REGION Network 157: Update the DAC for adjusting the VG2 voltage
   RUNG wire#powerrail
      { S7_Templates := "SrcType := Int" } LE_Contact(in1 := "STATO".stato_VOLTAGGIO_G2, in2 := 1150)
      { S7_Templates := "[SrcType := Int, DestType := Real]" } Convert(in := "STATO".stato_VOLTAGGIO_G2, out => "STATO_TMP".tmp_real_VG2)
      { S7_Templates := "SrcType := Real" } Mul(in1 := "STATO_TMP".tmp_real_VG2, in2 := 21.55, out => "STATO_TMP".tmp_real_VG2)
      { S7_Templates := "[SrcType := Real, DestType := DInt]" } Convert(in := "STATO_TMP".tmp_real_VG2, out => "STATO_TMP".tmp_adj_G2)
      { S7_Templates := "SrcType := DInt" } Mul(in1 := "STATO_TMP".tmp_adj_G2, in2 := "STATO".stato_adj_VG2, out => "STATO_TMP".tmp_adj_G2)
      { S7_Templates := "SrcType := DInt" } Div(in1 := "STATO_TMP".tmp_adj_G2, in2 := 1000, out => "dac_out_VG2")
   END_RUNG
   // the same network as SCL:
   IF "STATO".stato_VOLTAGGIO_G2 <= 1150 THEN
       "STATO_TMP".tmp_real_VG2 := INT_TO_REAL("STATO".stato_VOLTAGGIO_G2);
       "STATO_TMP".tmp_real_VG2 := "STATO_TMP".tmp_real_VG2 * 21.55;
       "STATO_TMP".tmp_adj_G2 := REAL_TO_DINT("STATO_TMP".tmp_real_VG2);
       "STATO_TMP".tmp_adj_G2 := "STATO_TMP".tmp_adj_G2 * "STATO".stato_adj_VG2;
       "dac_out_VG2" := "STATO_TMP".tmp_adj_G2 / 1000;
   END_IF;
END_REGION

REGION Network 158: Update the DAC for adjusting the VF voltage
   RUNG wire#powerrail
      { S7_Templates := "SrcType := Int" } LE_Contact(in1 := "STATO".stato_VOLTAGGIO_FILAMENTO, in2 := 8500)
      { S7_Templates := "[SrcType := Int, DestType := Real]" } Convert(in := "STATO".stato_VOLTAGGIO_FILAMENTO, out => "STATO_TMP".tmp_VFr)
      { S7_Templates := "SrcType := Real" } Div(in1 := "STATO_TMP".tmp_VFr, in2 := 1.0869, out => "STATO_TMP".tmp_VFr)
      { S7_Templates := "[SrcType := Real, DestType := Int]" } Convert(in := "STATO_TMP".tmp_VFr, out => "STATO_TMP".tmpVFi)
      { S7_Templates := "SrcType := DInt" } Mul(in1 := "STATO_TMP".tmpVFi, in2 := "STATO".stato_adj_VF, out => "STATO_TMP".tmp_adj_VF)
      { S7_Templates := "SrcType := DInt" } Div(in1 := "STATO_TMP".tmp_adj_VF, in2 := 1000, out => #dac_VF)
   END_RUNG
   // the same network as SCL:
   IF "STATO".stato_VOLTAGGIO_FILAMENTO <= 8500 THEN
       "STATO_TMP".tmp_VFr := INT_TO_REAL("STATO".stato_VOLTAGGIO_FILAMENTO);
       "STATO_TMP".tmp_VFr := "STATO_TMP".tmp_VFr / 1.0869;
       "STATO_TMP".tmpVFi := REAL_TO_INT("STATO_TMP".tmp_VFr);
       "STATO_TMP".tmp_adj_VF := "STATO_TMP".tmpVFi * "STATO".stato_adj_VF;
       #dac_VF := "STATO_TMP".tmp_adj_VF / 1000;
   END_IF;
END_REGION

REGION Network 159: Update the DAC for adjusting the VA voltage in CW
   // The voltage value must be below the threshold for CW mode.
   RUNG wire#powerrail
      Contact( "STATO".stato_MODO_CW )
      { S7_Templates := "SrcType := Int" } LE_Contact(in1 := "STATO".stato_ADJ_ANODICA_CW, in2 := "STATO".SOGLIA_VAcw)
      "REGOLA_ANODICA"(livello := "STATO".stato_ADJ_ANODICA_CW, uscita_dac => "dac_out_VA")
   END_RUNG
   // the same network as SCL:
   IF "STATO".stato_MODO_CW AND ("STATO".stato_ADJ_ANODICA_CW <= "STATO".SOGLIA_VAcw) THEN
       "REGOLA_ANODICA"(livello := "STATO".stato_ADJ_ANODICA_CW, uscita_dac => "dac_out_VA");
   END_IF;
END_REGION

REGION Network 160: Update the DAC for adjusting the VA voltage in Pulsed
   RUNG wire#powerrail
      Contact( "STATO".stato_MODO_PULSED )
      { S7_Templates := "SrcType := Int" } LE_Contact(in1 := "STATO".stato_ADJ_ANODICA_PULSED, in2 := 18000)
      "REGOLA_ANODICA"(livello := "STATO".stato_ADJ_ANODICA_PULSED, uscita_dac => "dac_out_VA")
   END_RUNG
   // the same network as SCL:
   IF "STATO".stato_MODO_PULSED AND ("STATO".stato_ADJ_ANODICA_PULSED <= 18000) THEN
       "REGOLA_ANODICA"(livello := "STATO".stato_ADJ_ANODICA_PULSED, uscita_dac => "dac_out_VA");
   END_IF;
END_REGION

REGION Network 161: Update the Reduced level
   RUNG wire#powerrail
      Contact( "STATO".controllo_setReduced )
      { S7_Templates := "SrcType := ???" } Mul(in1 := "STATO_TMP".tmp_Reduced, in2 := 10, out => "STATO".SogliaRidotta)
      Move(in := "STATO_TMP".tmp_Reduced, out1 => "STATO".stato_sogliaRIDOTTA)
      R_Coil( "STATO".controllo_setReduced )
   END_RUNG
   // the same network as SCL:
   IF "STATO".controllo_setReduced THEN
       "STATO".SogliaRidotta := "STATO_TMP".tmp_Reduced * 10;
       "STATO".stato_sogliaRIDOTTA := "STATO_TMP".tmp_Reduced;
       "STATO".controllo_setReduced := FALSE;
   END_IF;
END_REGION

REGION Network 162: Update the power levels for display panel
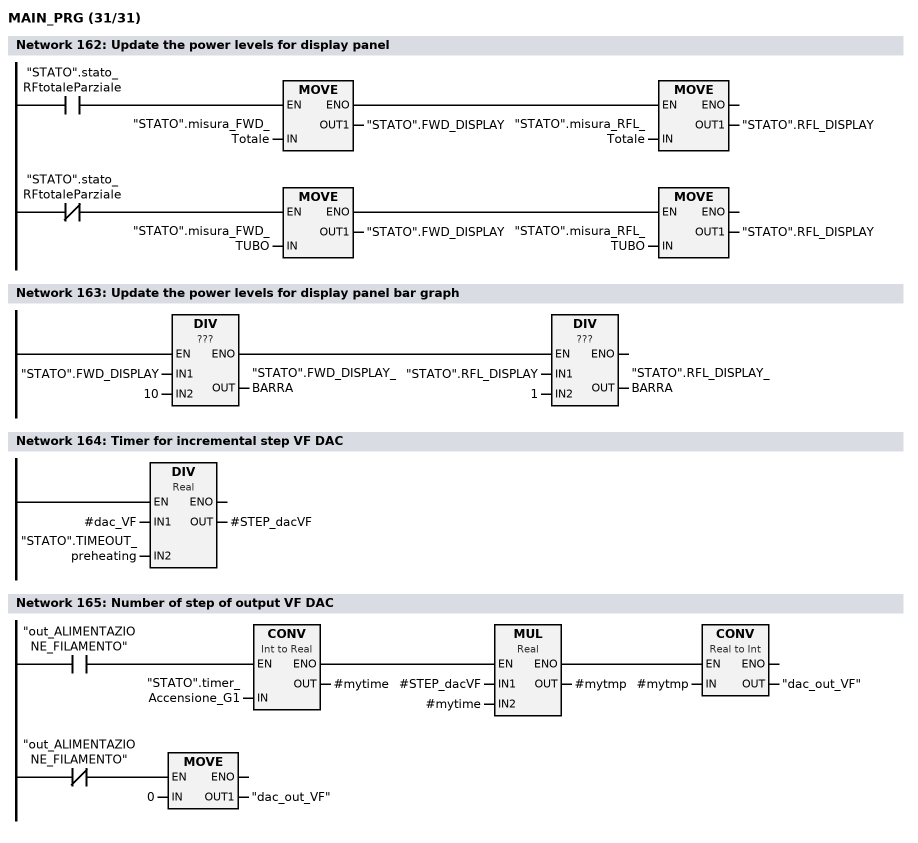
   RUNG wire#powerrail
      Contact( "STATO".stato_RFtotaleParziale )
      Move(in := "STATO".misura_FWD_Totale, out1 => "STATO".FWD_DISPLAY)
      Move(in := "STATO".misura_RFL_Totale, out1 => "STATO".RFL_DISPLAY)
   END_RUNG
   RUNG wire#powerrail
      I_Contact( "STATO".stato_RFtotaleParziale )
      Move(in := "STATO".misura_FWD_TUBO, out1 => "STATO".FWD_DISPLAY)
      Move(in := "STATO".misura_RFL_TUBO, out1 => "STATO".RFL_DISPLAY)
   END_RUNG
   // the same network as SCL:
   IF "STATO".stato_RFtotaleParziale THEN
       "STATO".FWD_DISPLAY := "STATO".misura_FWD_Totale;
       "STATO".RFL_DISPLAY := "STATO".misura_RFL_Totale;
   END_IF;
   IF NOT "STATO".stato_RFtotaleParziale THEN
       "STATO".FWD_DISPLAY := "STATO".misura_FWD_TUBO;
       "STATO".RFL_DISPLAY := "STATO".misura_RFL_TUBO;
   END_IF;
END_REGION

REGION Network 163: Update the power levels for display panel bar graph
   RUNG wire#powerrail
      { S7_Templates := "SrcType := ???" } Div(in1 := "STATO".FWD_DISPLAY, in2 := 10, out => "STATO".FWD_DISPLAY_BARRA)
      { S7_Templates := "SrcType := ???" } Div(in1 := "STATO".RFL_DISPLAY, in2 := 1, out => "STATO".RFL_DISPLAY_BARRA)
   END_RUNG
   // the same network as SCL:
   "STATO".FWD_DISPLAY_BARRA := "STATO".FWD_DISPLAY / 10;
   "STATO".RFL_DISPLAY_BARRA := "STATO".RFL_DISPLAY / 1;
END_REGION

REGION Network 164: Timer for incremental step VF DAC
   RUNG wire#powerrail
      { S7_Templates := "SrcType := Real" } Div(in1 := #dac_VF, in2 := "STATO".TIMEOUT_preheating, out => #STEP_dacVF)
   END_RUNG
   // the same network as SCL:
   #STEP_dacVF := #dac_VF / "STATO".TIMEOUT_preheating;
END_REGION

REGION Network 165: Number of step of output VF DAC
   RUNG wire#powerrail
      Contact( "out_ALIMENTAZIONE_FILAMENTO" )
      { S7_Templates := "[SrcType := Int, DestType := Real]" } Convert(in := "STATO".timer_Accensione_G1, out => #mytime)
      { S7_Templates := "SrcType := Real" } Mul(in1 := #STEP_dacVF, in2 := #mytime, out => #mytmp)
      { S7_Templates := "[SrcType := Real, DestType := Int]" } Convert(in := #mytmp, out => "dac_out_VF")
   END_RUNG
   RUNG wire#powerrail
      I_Contact( "out_ALIMENTAZIONE_FILAMENTO" )
      Move(in := 0, out1 => "dac_out_VF")
   END_RUNG
   // the same network as SCL:
   IF "out_ALIMENTAZIONE_FILAMENTO" THEN
       #mytime := INT_TO_REAL("STATO".timer_Accensione_G1);
       #mytmp := #STEP_dacVF * #mytime;
       "dac_out_VF" := REAL_TO_INT(#mytmp);
   END_IF;
   IF NOT "out_ALIMENTAZIONE_FILAMENTO" THEN "dac_out_VF" := 0; END_IF;
END_REGION
END_FUNCTION_BLOCK

FUNCTION "MISURE_ANALOGICHE" : Void   // FC1, LAD
TITLE = LETTURE ANALOGICHE DALL'ADC E DAL FLUSSOMETRO
{ S7_Optimized_Access := 'FALSE' }
VERSION : 0.1
   VAR_TEMP   // added for the SCL form of the ladder/FBD networks
      _w1 : Bool;
      _w2 : Bool;
      _w3 : Bool;
   END_VAR
BEGIN

REGION Network 1: MISURA TEMPERATURA LQD IN SS (1) bloccato
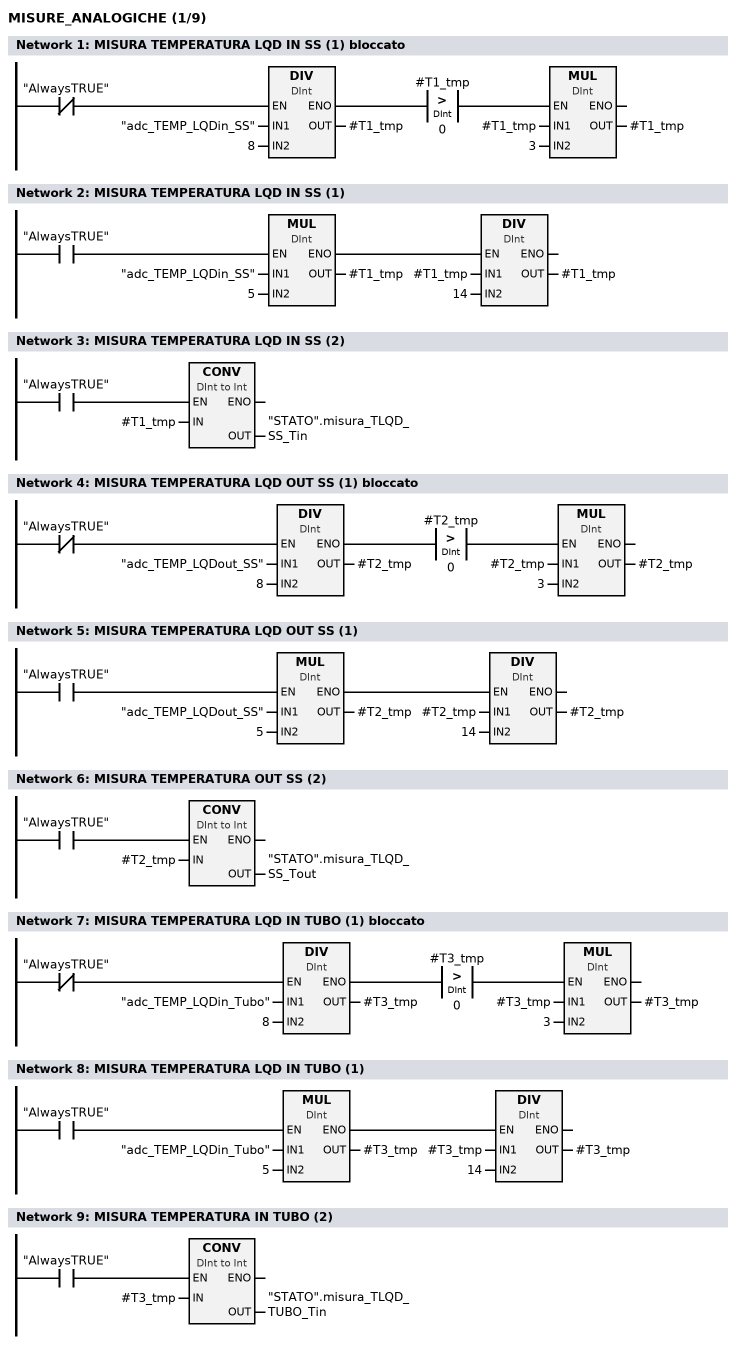
   RUNG wire#powerrail
      I_Contact( "AlwaysTRUE" )
      { S7_Templates := "SrcType := DInt" } Div(in1 := "adc_TEMP_LQDin_SS", in2 := 8, out => #T1_tmp)
      { S7_Templates := "SrcType := DInt" } GT_Contact(in1 := #T1_tmp, in2 := 0)
      { S7_Templates := "SrcType := DInt" } Mul(in1 := #T1_tmp, in2 := 3, out => #T1_tmp)
   END_RUNG
   // the same network as SCL:
   IF NOT "AlwaysTRUE" THEN #T1_tmp := "adc_TEMP_LQDin_SS" / 8; END_IF;
   IF NOT "AlwaysTRUE" AND (#T1_tmp > 0) THEN #T1_tmp := #T1_tmp * 3; END_IF;
END_REGION

REGION Network 2: MISURA TEMPERATURA LQD IN SS (1)
   RUNG wire#powerrail
      Contact( "AlwaysTRUE" )
      { S7_Templates := "SrcType := DInt" } Mul(in1 := "adc_TEMP_LQDin_SS", in2 := 5, out => #T1_tmp)
      { S7_Templates := "SrcType := DInt" } Div(in1 := #T1_tmp, in2 := 14, out => #T1_tmp)
   END_RUNG
   // the same network as SCL:
   IF "AlwaysTRUE" THEN
       #T1_tmp := "adc_TEMP_LQDin_SS" * 5;
       #T1_tmp := #T1_tmp / 14;
   END_IF;
END_REGION

REGION Network 3: MISURA TEMPERATURA LQD IN SS (2)
   RUNG wire#powerrail
      Contact( "AlwaysTRUE" )
      { S7_Templates := "[SrcType := DInt, DestType := Int]" } Convert(in := #T1_tmp, out => "STATO".misura_TLQD_SS_Tin)
   END_RUNG
   // the same network as SCL:
   IF "AlwaysTRUE" THEN "STATO".misura_TLQD_SS_Tin := DINT_TO_INT(#T1_tmp); END_IF;
END_REGION

REGION Network 4: MISURA TEMPERATURA LQD OUT SS (1) bloccato
   RUNG wire#powerrail
      I_Contact( "AlwaysTRUE" )
      { S7_Templates := "SrcType := DInt" } Div(in1 := "adc_TEMP_LQDout_SS", in2 := 8, out => #T2_tmp)
      { S7_Templates := "SrcType := DInt" } GT_Contact(in1 := #T2_tmp, in2 := 0)
      { S7_Templates := "SrcType := DInt" } Mul(in1 := #T2_tmp, in2 := 3, out => #T2_tmp)
   END_RUNG
   // the same network as SCL:
   IF NOT "AlwaysTRUE" THEN #T2_tmp := "adc_TEMP_LQDout_SS" / 8; END_IF;
   IF NOT "AlwaysTRUE" AND (#T2_tmp > 0) THEN #T2_tmp := #T2_tmp * 3; END_IF;
END_REGION

REGION Network 5: MISURA TEMPERATURA LQD OUT SS (1)
   RUNG wire#powerrail
      Contact( "AlwaysTRUE" )
      { S7_Templates := "SrcType := DInt" } Mul(in1 := "adc_TEMP_LQDout_SS", in2 := 5, out => #T2_tmp)
      { S7_Templates := "SrcType := DInt" } Div(in1 := #T2_tmp, in2 := 14, out => #T2_tmp)
   END_RUNG
   // the same network as SCL:
   IF "AlwaysTRUE" THEN
       #T2_tmp := "adc_TEMP_LQDout_SS" * 5;
       #T2_tmp := #T2_tmp / 14;
   END_IF;
END_REGION

REGION Network 6: MISURA TEMPERATURA OUT SS (2)
   RUNG wire#powerrail
      Contact( "AlwaysTRUE" )
      { S7_Templates := "[SrcType := DInt, DestType := Int]" } Convert(in := #T2_tmp, out => "STATO".misura_TLQD_SS_Tout)
   END_RUNG
   // the same network as SCL:
   IF "AlwaysTRUE" THEN "STATO".misura_TLQD_SS_Tout := DINT_TO_INT(#T2_tmp); END_IF;
END_REGION

REGION Network 7: MISURA TEMPERATURA LQD IN TUBO (1) bloccato
   RUNG wire#powerrail
      I_Contact( "AlwaysTRUE" )
      { S7_Templates := "SrcType := DInt" } Div(in1 := "adc_TEMP_LQDin_Tubo", in2 := 8, out => #T3_tmp)
      { S7_Templates := "SrcType := DInt" } GT_Contact(in1 := #T3_tmp, in2 := 0)
      { S7_Templates := "SrcType := DInt" } Mul(in1 := #T3_tmp, in2 := 3, out => #T3_tmp)
   END_RUNG
   // the same network as SCL:
   IF NOT "AlwaysTRUE" THEN #T3_tmp := "adc_TEMP_LQDin_Tubo" / 8; END_IF;
   IF NOT "AlwaysTRUE" AND (#T3_tmp > 0) THEN #T3_tmp := #T3_tmp * 3; END_IF;
END_REGION

REGION Network 8: MISURA TEMPERATURA LQD IN TUBO (1)
   RUNG wire#powerrail
      Contact( "AlwaysTRUE" )
      { S7_Templates := "SrcType := DInt" } Mul(in1 := "adc_TEMP_LQDin_Tubo", in2 := 5, out => #T3_tmp)
      { S7_Templates := "SrcType := DInt" } Div(in1 := #T3_tmp, in2 := 14, out => #T3_tmp)
   END_RUNG
   // the same network as SCL:
   IF "AlwaysTRUE" THEN
       #T3_tmp := "adc_TEMP_LQDin_Tubo" * 5;
       #T3_tmp := #T3_tmp / 14;
   END_IF;
END_REGION

REGION Network 9: MISURA TEMPERATURA IN TUBO (2)
   RUNG wire#powerrail
      Contact( "AlwaysTRUE" )
      { S7_Templates := "[SrcType := DInt, DestType := Int]" } Convert(in := #T3_tmp, out => "STATO".misura_TLQD_TUBO_Tin)
   END_RUNG
   // the same network as SCL:
   IF "AlwaysTRUE" THEN "STATO".misura_TLQD_TUBO_Tin := DINT_TO_INT(#T3_tmp); END_IF;
END_REGION

REGION Network 10: MISURA TEMPERATURA LQD OUT TUBO (1) bloccato
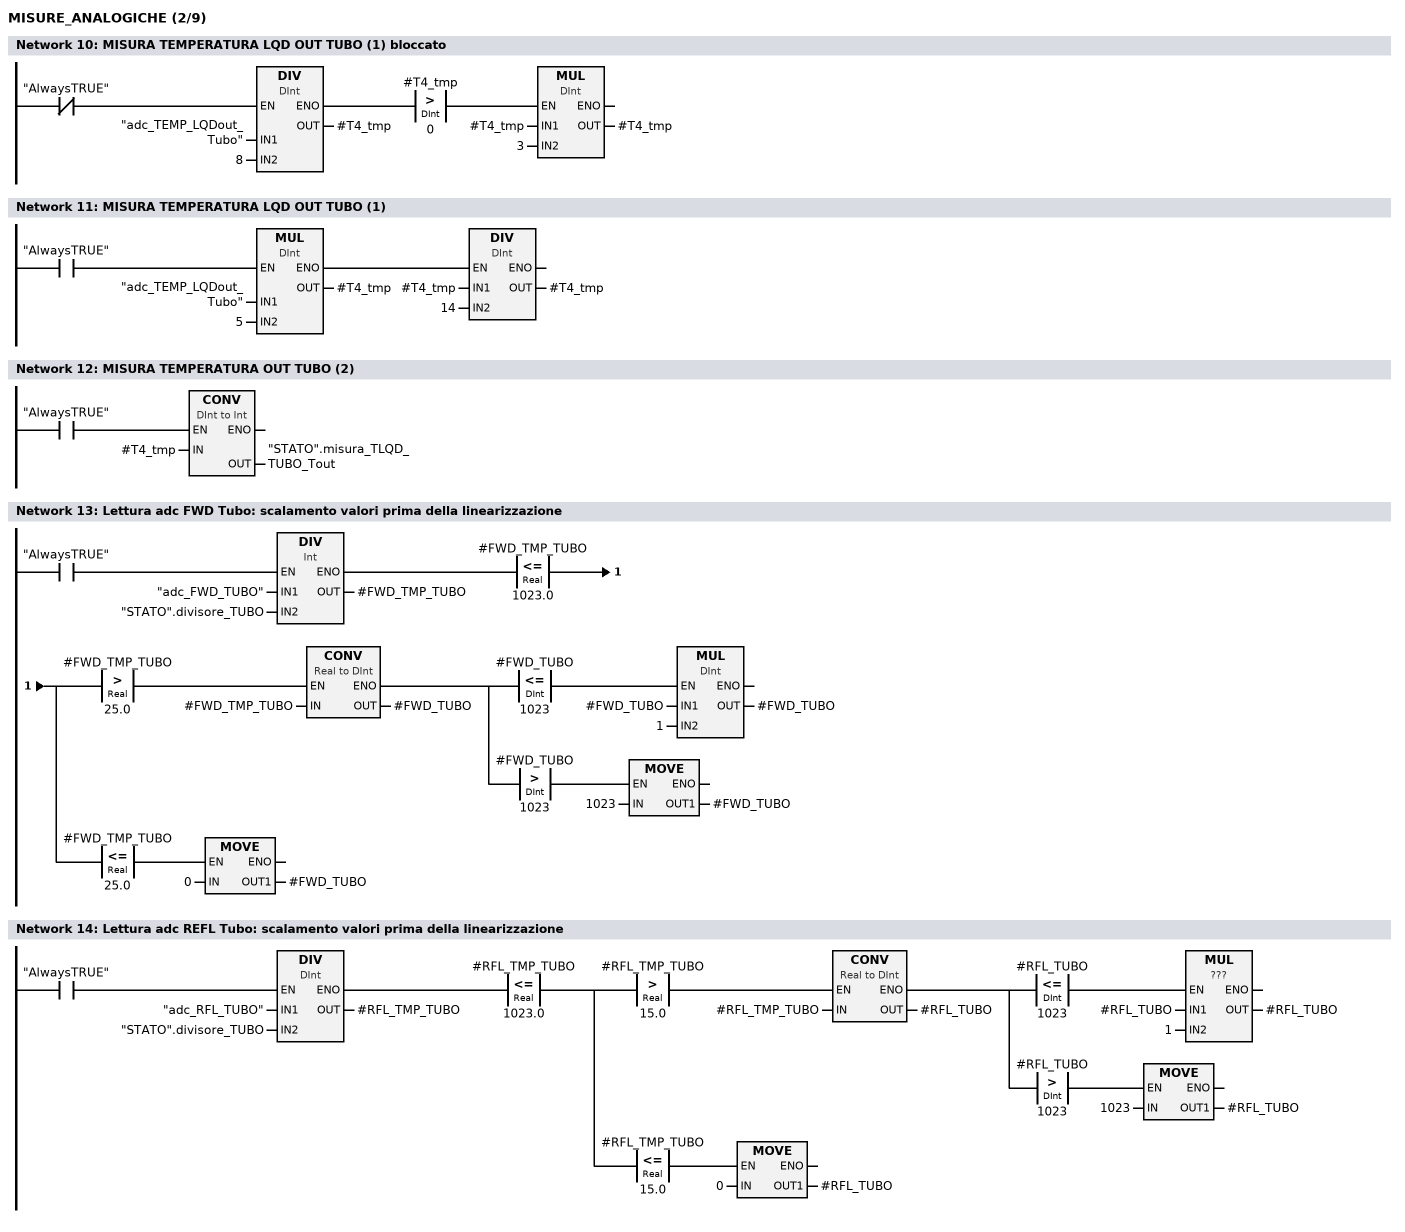
   RUNG wire#powerrail
      I_Contact( "AlwaysTRUE" )
      { S7_Templates := "SrcType := DInt" } Div(in1 := "adc_TEMP_LQDout_Tubo", in2 := 8, out => #T4_tmp)
      { S7_Templates := "SrcType := DInt" } GT_Contact(in1 := #T4_tmp, in2 := 0)
      { S7_Templates := "SrcType := DInt" } Mul(in1 := #T4_tmp, in2 := 3, out => #T4_tmp)
   END_RUNG
   // the same network as SCL:
   IF NOT "AlwaysTRUE" THEN #T4_tmp := "adc_TEMP_LQDout_Tubo" / 8; END_IF;
   IF NOT "AlwaysTRUE" AND (#T4_tmp > 0) THEN #T4_tmp := #T4_tmp * 3; END_IF;
END_REGION

REGION Network 11: MISURA TEMPERATURA LQD OUT TUBO (1)
   RUNG wire#powerrail
      Contact( "AlwaysTRUE" )
      { S7_Templates := "SrcType := DInt" } Mul(in1 := "adc_TEMP_LQDout_Tubo", in2 := 5, out => #T4_tmp)
      { S7_Templates := "SrcType := DInt" } Div(in1 := #T4_tmp, in2 := 14, out => #T4_tmp)
   END_RUNG
   // the same network as SCL:
   IF "AlwaysTRUE" THEN
       #T4_tmp := "adc_TEMP_LQDout_Tubo" * 5;
       #T4_tmp := #T4_tmp / 14;
   END_IF;
END_REGION

REGION Network 12: MISURA TEMPERATURA OUT TUBO (2)
   RUNG wire#powerrail
      Contact( "AlwaysTRUE" )
      { S7_Templates := "[SrcType := DInt, DestType := Int]" } Convert(in := #T4_tmp, out => "STATO".misura_TLQD_TUBO_Tout)
   END_RUNG
   // the same network as SCL:
   IF "AlwaysTRUE" THEN "STATO".misura_TLQD_TUBO_Tout := DINT_TO_INT(#T4_tmp); END_IF;
END_REGION

REGION Network 13: Lettura adc FWD Tubo: scalamento valori prima della linearizzazione
   RUNG wire#powerrail
      Contact( "AlwaysTRUE" )
      { S7_Templates := "SrcType := Int" } Div(in1 := "adc_FWD_TUBO", in2 := "STATO".divisore_TUBO, out => #FWD_TMP_TUBO)
      { S7_Templates := "SrcType := Real" } LE_Contact(in1 := #FWD_TMP_TUBO, in2 := 1023.0)
      wire#w1
      { S7_Templates := "SrcType := Real" } GT_Contact(in1 := #FWD_TMP_TUBO, in2 := 25.0)
      { S7_Templates := "[SrcType := Real, DestType := DInt]" } Convert(in := #FWD_TMP_TUBO, out => #FWD_TUBO)
      wire#w2
      { S7_Templates := "SrcType := DInt" } LE_Contact(in1 := #FWD_TUBO, in2 := 1023)
      { S7_Templates := "SrcType := DInt" } Mul(in1 := #FWD_TUBO, in2 := 1, out => #FWD_TUBO)
   END_RUNG
   RUNG wire#w2
      { S7_Templates := "SrcType := DInt" } GT_Contact(in1 := #FWD_TUBO, in2 := 1023)
      Move(in := 1023, out1 => #FWD_TUBO)
   END_RUNG
   RUNG wire#w1
      { S7_Templates := "SrcType := Real" } LE_Contact(in1 := #FWD_TMP_TUBO, in2 := 25.0)
      Move(in := 0, out1 => #FWD_TUBO)
   END_RUNG
   // the same network as SCL:
   IF "AlwaysTRUE" THEN #FWD_TMP_TUBO := "adc_FWD_TUBO" / "STATO".divisore_TUBO; END_IF;
   #_w1 := "AlwaysTRUE" AND (#FWD_TMP_TUBO <= 1023.0);
   #_w2 := #_w1 AND (#FWD_TMP_TUBO > 25.0);
   IF #_w2 THEN #FWD_TUBO := REAL_TO_DINT(#FWD_TMP_TUBO); END_IF;
   IF #_w2 AND (#FWD_TUBO <= 1023) THEN #FWD_TUBO := #FWD_TUBO * 1; END_IF;
   IF #_w2 AND (#FWD_TUBO > 1023) THEN #FWD_TUBO := 1023; END_IF;
   IF #_w1 AND (#FWD_TMP_TUBO <= 25.0) THEN #FWD_TUBO := 0; END_IF;
END_REGION

REGION Network 14: Lettura adc REFL Tubo: scalamento valori prima della linearizzazione
   RUNG wire#powerrail
      Contact( "AlwaysTRUE" )
      { S7_Templates := "SrcType := DInt" } Div(in1 := "adc_RFL_TUBO", in2 := "STATO".divisore_TUBO, out => #RFL_TMP_TUBO)
      { S7_Templates := "SrcType := Real" } LE_Contact(in1 := #RFL_TMP_TUBO, in2 := 1023.0)
      wire#w1
      { S7_Templates := "SrcType := Real" } GT_Contact(in1 := #RFL_TMP_TUBO, in2 := 15.0)
      { S7_Templates := "[SrcType := Real, DestType := DInt]" } Convert(in := #RFL_TMP_TUBO, out => #RFL_TUBO)
      wire#w2
      { S7_Templates := "SrcType := DInt" } LE_Contact(in1 := #RFL_TUBO, in2 := 1023)
      { S7_Templates := "SrcType := ???" } Mul(in1 := #RFL_TUBO, in2 := 1, out => #RFL_TUBO)
   END_RUNG
   RUNG wire#w2
      { S7_Templates := "SrcType := DInt" } GT_Contact(in1 := #RFL_TUBO, in2 := 1023)
      Move(in := 1023, out1 => #RFL_TUBO)
   END_RUNG
   RUNG wire#w1
      { S7_Templates := "SrcType := Real" } LE_Contact(in1 := #RFL_TMP_TUBO, in2 := 15.0)
      Move(in := 0, out1 => #RFL_TUBO)
   END_RUNG
   // the same network as SCL:
   IF "AlwaysTRUE" THEN #RFL_TMP_TUBO := "adc_RFL_TUBO" / "STATO".divisore_TUBO; END_IF;
   #_w1 := "AlwaysTRUE" AND (#RFL_TMP_TUBO <= 1023.0);
   #_w2 := #_w1 AND (#RFL_TMP_TUBO > 15.0);
   IF #_w2 THEN #RFL_TUBO := REAL_TO_DINT(#RFL_TMP_TUBO); END_IF;
   IF #_w2 AND (#RFL_TUBO <= 1023) THEN #RFL_TUBO := #RFL_TUBO * 1; END_IF;
   IF #_w2 AND (#RFL_TUBO > 1023) THEN #RFL_TUBO := 1023; END_IF;
   IF #_w1 AND (#RFL_TMP_TUBO <= 15.0) THEN #RFL_TUBO := 0; END_IF;
END_REGION

REGION Network 15: Lettura adc FWD Stato Solido: scalamento valori prima della linearizzazione
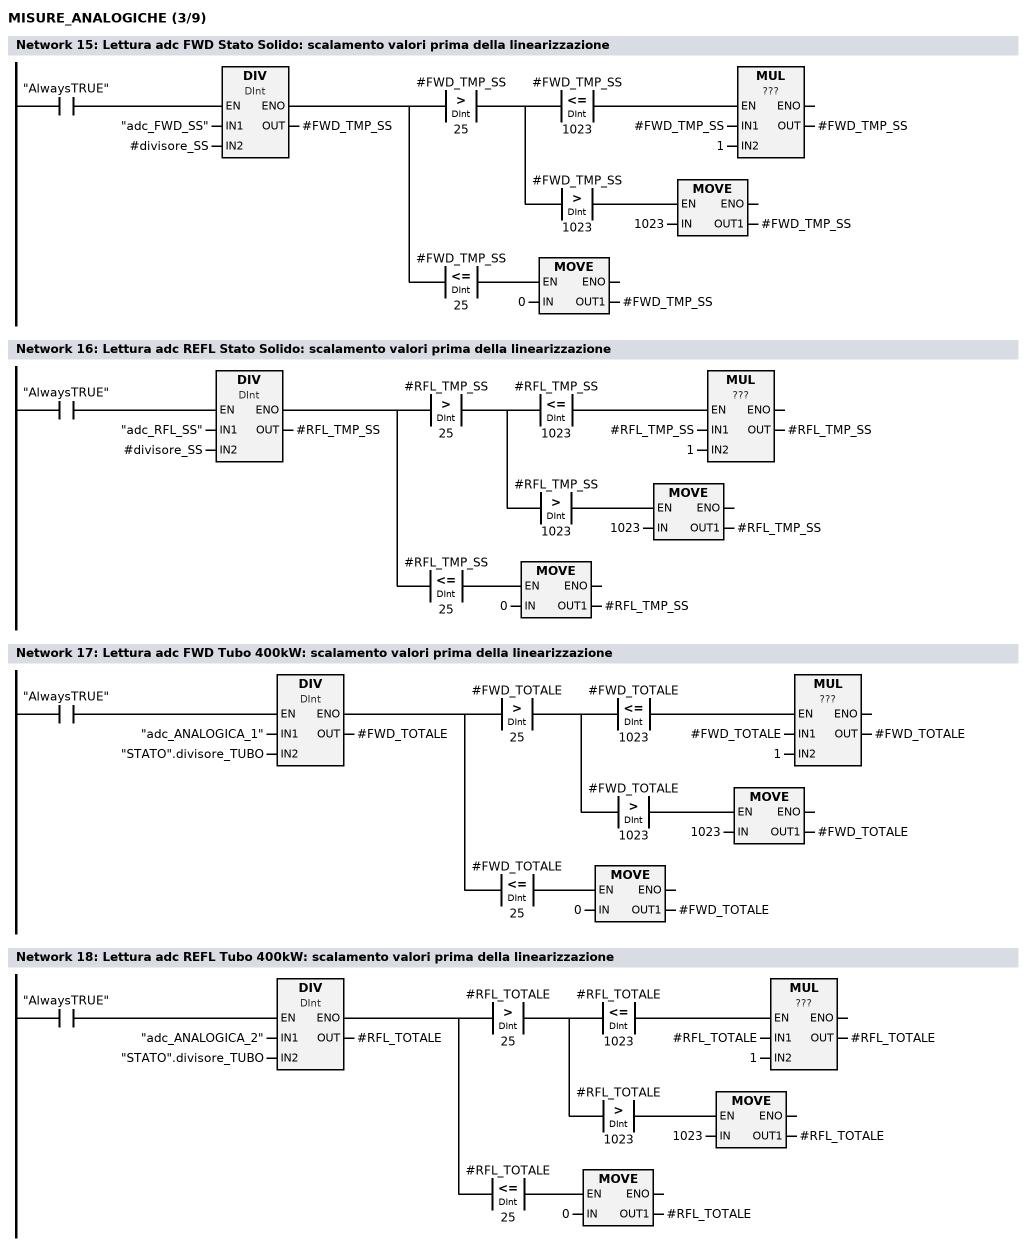
   RUNG wire#powerrail
      Contact( "AlwaysTRUE" )
      { S7_Templates := "SrcType := DInt" } Div(in1 := "adc_FWD_SS", in2 := #divisore_SS, out => #FWD_TMP_SS)
      wire#w1
      { S7_Templates := "SrcType := DInt" } GT_Contact(in1 := #FWD_TMP_SS, in2 := 25)
      wire#w2
      { S7_Templates := "SrcType := DInt" } LE_Contact(in1 := #FWD_TMP_SS, in2 := 1023)
      { S7_Templates := "SrcType := ???" } Mul(in1 := #FWD_TMP_SS, in2 := 1, out => #FWD_TMP_SS)
   END_RUNG
   RUNG wire#w2
      { S7_Templates := "SrcType := DInt" } GT_Contact(in1 := #FWD_TMP_SS, in2 := 1023)
      Move(in := 1023, out1 => #FWD_TMP_SS)
   END_RUNG
   RUNG wire#w1
      { S7_Templates := "SrcType := DInt" } LE_Contact(in1 := #FWD_TMP_SS, in2 := 25)
      Move(in := 0, out1 => #FWD_TMP_SS)
   END_RUNG
   // the same network as SCL:
   IF "AlwaysTRUE" THEN #FWD_TMP_SS := "adc_FWD_SS" / #divisore_SS; END_IF;
   #_w1 := "AlwaysTRUE" AND (#FWD_TMP_SS > 25);
   IF #_w1 AND (#FWD_TMP_SS <= 1023) THEN #FWD_TMP_SS := #FWD_TMP_SS * 1; END_IF;
   IF #_w1 AND (#FWD_TMP_SS > 1023) THEN #FWD_TMP_SS := 1023; END_IF;
   IF "AlwaysTRUE" AND (#FWD_TMP_SS <= 25) THEN #FWD_TMP_SS := 0; END_IF;
END_REGION

REGION Network 16: Lettura adc REFL Stato Solido: scalamento valori prima della linearizzazione
   RUNG wire#powerrail
      Contact( "AlwaysTRUE" )
      { S7_Templates := "SrcType := DInt" } Div(in1 := "adc_RFL_SS", in2 := #divisore_SS, out => #RFL_TMP_SS)
      wire#w1
      { S7_Templates := "SrcType := DInt" } GT_Contact(in1 := #RFL_TMP_SS, in2 := 25)
      wire#w2
      { S7_Templates := "SrcType := DInt" } LE_Contact(in1 := #RFL_TMP_SS, in2 := 1023)
      { S7_Templates := "SrcType := ???" } Mul(in1 := #RFL_TMP_SS, in2 := 1, out => #RFL_TMP_SS)
   END_RUNG
   RUNG wire#w2
      { S7_Templates := "SrcType := DInt" } GT_Contact(in1 := #RFL_TMP_SS, in2 := 1023)
      Move(in := 1023, out1 => #RFL_TMP_SS)
   END_RUNG
   RUNG wire#w1
      { S7_Templates := "SrcType := DInt" } LE_Contact(in1 := #RFL_TMP_SS, in2 := 25)
      Move(in := 0, out1 => #RFL_TMP_SS)
   END_RUNG
   // the same network as SCL:
   IF "AlwaysTRUE" THEN #RFL_TMP_SS := "adc_RFL_SS" / #divisore_SS; END_IF;
   #_w1 := "AlwaysTRUE" AND (#RFL_TMP_SS > 25);
   IF #_w1 AND (#RFL_TMP_SS <= 1023) THEN #RFL_TMP_SS := #RFL_TMP_SS * 1; END_IF;
   IF #_w1 AND (#RFL_TMP_SS > 1023) THEN #RFL_TMP_SS := 1023; END_IF;
   IF "AlwaysTRUE" AND (#RFL_TMP_SS <= 25) THEN #RFL_TMP_SS := 0; END_IF;
END_REGION

REGION Network 17: Lettura adc FWD Tubo 400kW: scalamento valori prima della linearizzazione
   RUNG wire#powerrail
      Contact( "AlwaysTRUE" )
      { S7_Templates := "SrcType := DInt" } Div(in1 := "adc_ANALOGICA_1", in2 := "STATO".divisore_TUBO, out => #FWD_TOTALE)
      wire#w1
      { S7_Templates := "SrcType := DInt" } GT_Contact(in1 := #FWD_TOTALE, in2 := 25)
      wire#w2
      { S7_Templates := "SrcType := DInt" } LE_Contact(in1 := #FWD_TOTALE, in2 := 1023)
      { S7_Templates := "SrcType := ???" } Mul(in1 := #FWD_TOTALE, in2 := 1, out => #FWD_TOTALE)
   END_RUNG
   RUNG wire#w2
      { S7_Templates := "SrcType := DInt" } GT_Contact(in1 := #FWD_TOTALE, in2 := 1023)
      Move(in := 1023, out1 => #FWD_TOTALE)
   END_RUNG
   RUNG wire#w1
      { S7_Templates := "SrcType := DInt" } LE_Contact(in1 := #FWD_TOTALE, in2 := 25)
      Move(in := 0, out1 => #FWD_TOTALE)
   END_RUNG
   // the same network as SCL:
   IF "AlwaysTRUE" THEN #FWD_TOTALE := "adc_ANALOGICA_1" / "STATO".divisore_TUBO; END_IF;
   #_w1 := "AlwaysTRUE" AND (#FWD_TOTALE > 25);
   IF #_w1 AND (#FWD_TOTALE <= 1023) THEN #FWD_TOTALE := #FWD_TOTALE * 1; END_IF;
   IF #_w1 AND (#FWD_TOTALE > 1023) THEN #FWD_TOTALE := 1023; END_IF;
   IF "AlwaysTRUE" AND (#FWD_TOTALE <= 25) THEN #FWD_TOTALE := 0; END_IF;
END_REGION

REGION Network 18: Lettura adc REFL Tubo 400kW: scalamento valori prima della linearizzazione
   RUNG wire#powerrail
      Contact( "AlwaysTRUE" )
      { S7_Templates := "SrcType := DInt" } Div(in1 := "adc_ANALOGICA_2", in2 := "STATO".divisore_TUBO, out => #RFL_TOTALE)
      wire#w1
      { S7_Templates := "SrcType := DInt" } GT_Contact(in1 := #RFL_TOTALE, in2 := 25)
      wire#w2
      { S7_Templates := "SrcType := DInt" } LE_Contact(in1 := #RFL_TOTALE, in2 := 1023)
      { S7_Templates := "SrcType := ???" } Mul(in1 := #RFL_TOTALE, in2 := 1, out => #RFL_TOTALE)
   END_RUNG
   RUNG wire#w2
      { S7_Templates := "SrcType := DInt" } GT_Contact(in1 := #RFL_TOTALE, in2 := 1023)
      Move(in := 1023, out1 => #RFL_TOTALE)
   END_RUNG
   RUNG wire#w1
      { S7_Templates := "SrcType := DInt" } LE_Contact(in1 := #RFL_TOTALE, in2 := 25)
      Move(in := 0, out1 => #RFL_TOTALE)
   END_RUNG
   // the same network as SCL:
   IF "AlwaysTRUE" THEN #RFL_TOTALE := "adc_ANALOGICA_2" / "STATO".divisore_TUBO; END_IF;
   #_w1 := "AlwaysTRUE" AND (#RFL_TOTALE > 25);
   IF #_w1 AND (#RFL_TOTALE <= 1023) THEN #RFL_TOTALE := #RFL_TOTALE * 1; END_IF;
   IF #_w1 AND (#RFL_TOTALE > 1023) THEN #RFL_TOTALE := 1023; END_IF;
   IF "AlwaysTRUE" AND (#RFL_TOTALE <= 25) THEN #RFL_TOTALE := 0; END_IF;
END_REGION

REGION Network 19: Linearizzazione FWD Tubo 200kW
   // Impulsivo o CW
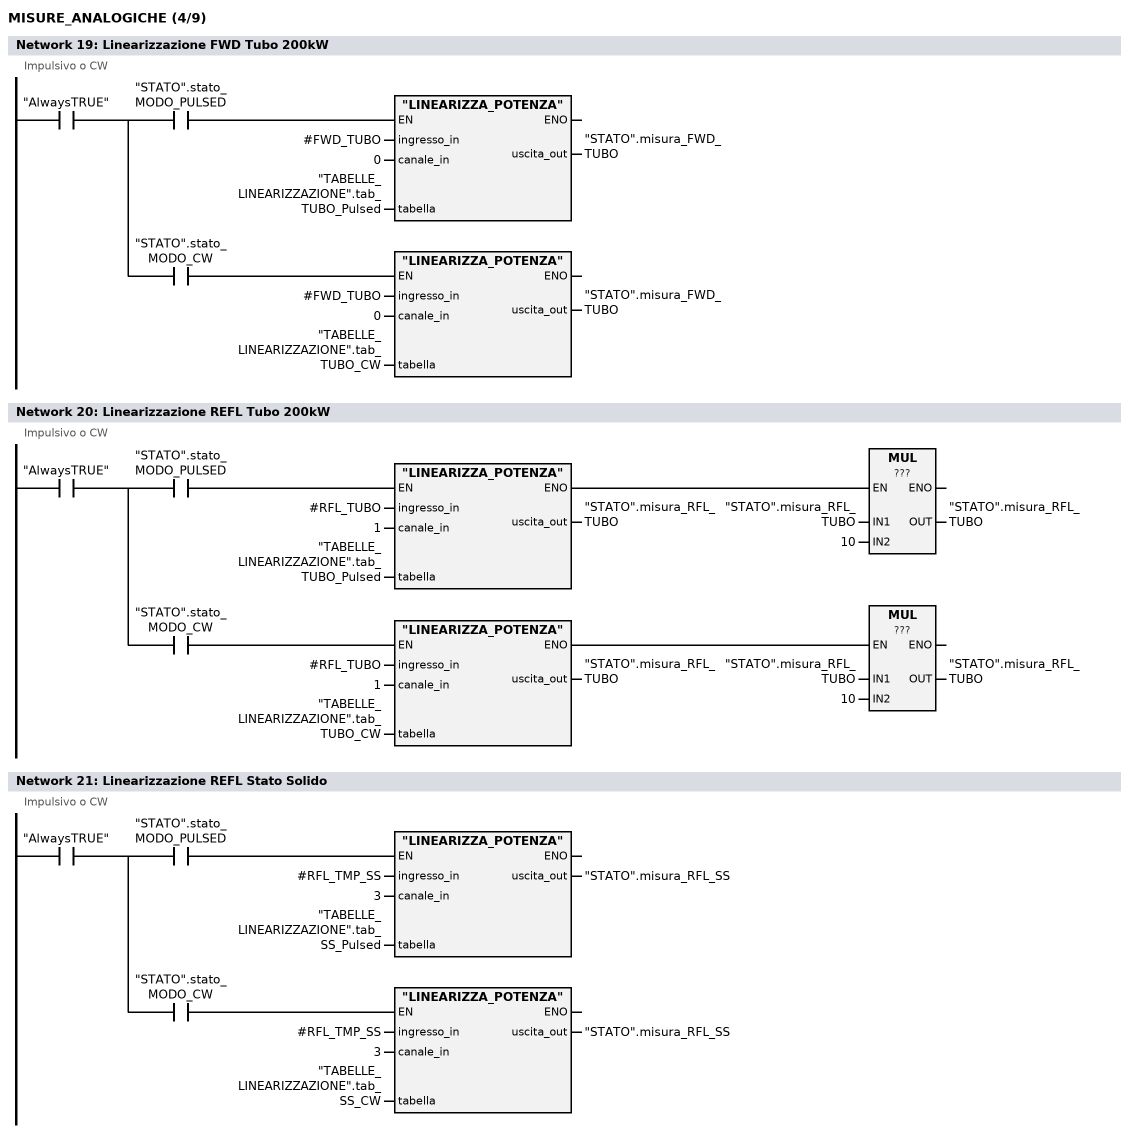
   RUNG wire#powerrail
      Contact( "AlwaysTRUE" )
      wire#w1
      Contact( "STATO".stato_MODO_PULSED )
      "LINEARIZZA_POTENZA"(ingresso_in := #FWD_TUBO, canale_in := 0, tabella := "TABELLE_LINEARIZZAZIONE".tab_TUBO_Pulsed, uscita_out => "STATO".misura_FWD_TUBO)
   END_RUNG
   RUNG wire#w1
      Contact( "STATO".stato_MODO_CW )
      "LINEARIZZA_POTENZA"(ingresso_in := #FWD_TUBO, canale_in := 0, tabella := "TABELLE_LINEARIZZAZIONE".tab_TUBO_CW, uscita_out => "STATO".misura_FWD_TUBO)
   END_RUNG
   // the same network as SCL:
   #_w1 := "AlwaysTRUE";
   IF "AlwaysTRUE" AND "STATO".stato_MODO_PULSED THEN
       "LINEARIZZA_POTENZA"(ingresso_in := #FWD_TUBO,
                            canale_in := 0,
                            tabella := "TABELLE_LINEARIZZAZIONE".tab_TUBO_Pulsed,
                            uscita_out => "STATO".misura_FWD_TUBO);
   END_IF;
   IF #_w1 AND "STATO".stato_MODO_CW THEN
       "LINEARIZZA_POTENZA"(ingresso_in := #FWD_TUBO,
                            canale_in := 0,
                            tabella := "TABELLE_LINEARIZZAZIONE".tab_TUBO_CW,
                            uscita_out => "STATO".misura_FWD_TUBO);
   END_IF;
END_REGION

REGION Network 20: Linearizzazione REFL Tubo 200kW
   // Impulsivo o CW
   RUNG wire#powerrail
      Contact( "AlwaysTRUE" )
      wire#w1
      Contact( "STATO".stato_MODO_PULSED )
      "LINEARIZZA_POTENZA"(ingresso_in := #RFL_TUBO, canale_in := 1, tabella := "TABELLE_LINEARIZZAZIONE".tab_TUBO_Pulsed, uscita_out => "STATO".misura_RFL_TUBO)
      { S7_Templates := "SrcType := ???" } Mul(in1 := "STATO".misura_RFL_TUBO, in2 := 10, out => "STATO".misura_RFL_TUBO)
   END_RUNG
   RUNG wire#w1
      Contact( "STATO".stato_MODO_CW )
      "LINEARIZZA_POTENZA"(ingresso_in := #RFL_TUBO, canale_in := 1, tabella := "TABELLE_LINEARIZZAZIONE".tab_TUBO_CW, uscita_out => "STATO".misura_RFL_TUBO)
      { S7_Templates := "SrcType := ???" } Mul(in1 := "STATO".misura_RFL_TUBO, in2 := 10, out => "STATO".misura_RFL_TUBO)
   END_RUNG
   // the same network as SCL:
   #_w2 := "AlwaysTRUE";
   "LINEARIZZA_POTENZA"(EN := "AlwaysTRUE" AND "STATO".stato_MODO_PULSED,
                        ingresso_in := #RFL_TUBO,
                        canale_in := 1,
                        tabella := "TABELLE_LINEARIZZAZIONE".tab_TUBO_Pulsed,
                        uscita_out => "STATO".misura_RFL_TUBO,
                        ENO => #_w1);
   IF #_w1 THEN "STATO".misura_RFL_TUBO := "STATO".misura_RFL_TUBO * 10; END_IF;
   "LINEARIZZA_POTENZA"(EN := #_w2 AND "STATO".stato_MODO_CW,
                        ingresso_in := #RFL_TUBO,
                        canale_in := 1,
                        tabella := "TABELLE_LINEARIZZAZIONE".tab_TUBO_CW,
                        uscita_out => "STATO".misura_RFL_TUBO,
                        ENO => #_w3);
   IF #_w3 THEN "STATO".misura_RFL_TUBO := "STATO".misura_RFL_TUBO * 10; END_IF;
END_REGION

REGION Network 21: Linearizzazione REFL Stato Solido
   // Impulsivo o CW
   RUNG wire#powerrail
      Contact( "AlwaysTRUE" )
      wire#w1
      Contact( "STATO".stato_MODO_PULSED )
      "LINEARIZZA_POTENZA"(ingresso_in := #RFL_TMP_SS, canale_in := 3, tabella := "TABELLE_LINEARIZZAZIONE".tab_SS_Pulsed, uscita_out => "STATO".misura_RFL_SS)
   END_RUNG
   RUNG wire#w1
      Contact( "STATO".stato_MODO_CW )
      "LINEARIZZA_POTENZA"(ingresso_in := #RFL_TMP_SS, canale_in := 3, tabella := "TABELLE_LINEARIZZAZIONE".tab_SS_CW, uscita_out => "STATO".misura_RFL_SS)
   END_RUNG
   // the same network as SCL:
   #_w1 := "AlwaysTRUE";
   IF "AlwaysTRUE" AND "STATO".stato_MODO_PULSED THEN
       "LINEARIZZA_POTENZA"(ingresso_in := #RFL_TMP_SS,
                            canale_in := 3,
                            tabella := "TABELLE_LINEARIZZAZIONE".tab_SS_Pulsed,
                            uscita_out => "STATO".misura_RFL_SS);
   END_IF;
   IF #_w1 AND "STATO".stato_MODO_CW THEN
       "LINEARIZZA_POTENZA"(ingresso_in := #RFL_TMP_SS,
                            canale_in := 3,
                            tabella := "TABELLE_LINEARIZZAZIONE".tab_SS_CW,
                            uscita_out => "STATO".misura_RFL_SS);
   END_IF;
END_REGION

REGION Network 22: Linearizzazione FWD Stato Solido
   // Impulsivo o CW
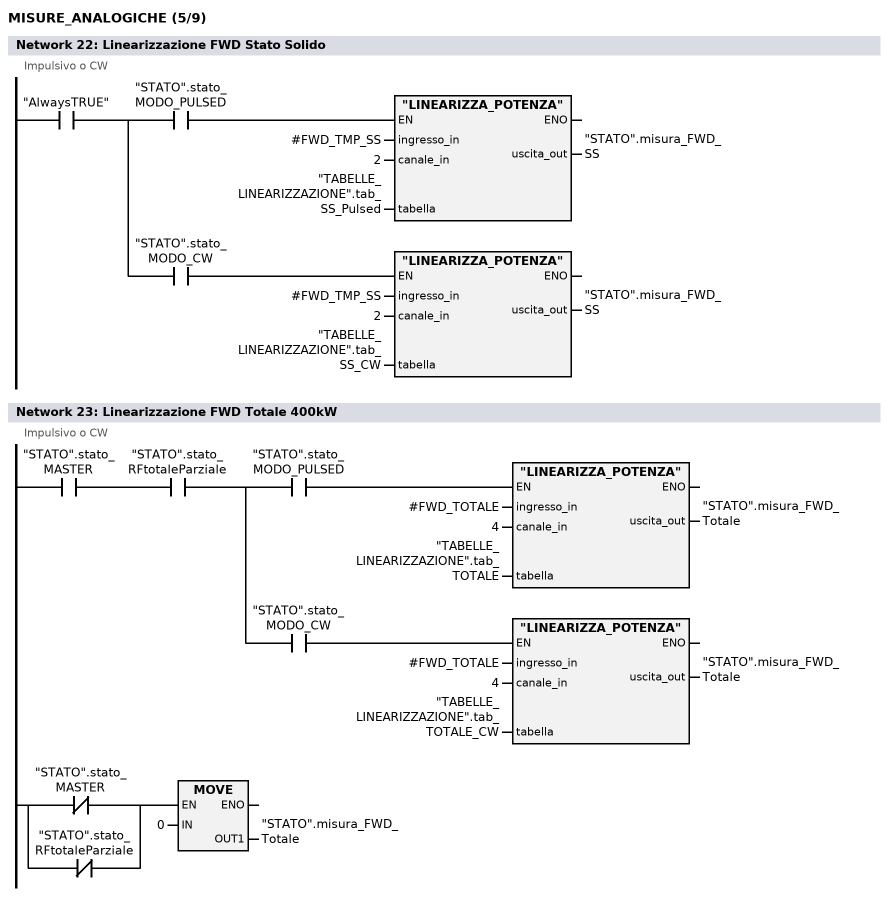
   RUNG wire#powerrail
      Contact( "AlwaysTRUE" )
      wire#w1
      Contact( "STATO".stato_MODO_PULSED )
      "LINEARIZZA_POTENZA"(ingresso_in := #FWD_TMP_SS, canale_in := 2, tabella := "TABELLE_LINEARIZZAZIONE".tab_SS_Pulsed, uscita_out => "STATO".misura_FWD_SS)
   END_RUNG
   RUNG wire#w1
      Contact( "STATO".stato_MODO_CW )
      "LINEARIZZA_POTENZA"(ingresso_in := #FWD_TMP_SS, canale_in := 2, tabella := "TABELLE_LINEARIZZAZIONE".tab_SS_CW, uscita_out => "STATO".misura_FWD_SS)
   END_RUNG
   // the same network as SCL:
   #_w1 := "AlwaysTRUE";
   IF "AlwaysTRUE" AND "STATO".stato_MODO_PULSED THEN
       "LINEARIZZA_POTENZA"(ingresso_in := #FWD_TMP_SS,
                            canale_in := 2,
                            tabella := "TABELLE_LINEARIZZAZIONE".tab_SS_Pulsed,
                            uscita_out => "STATO".misura_FWD_SS);
   END_IF;
   IF #_w1 AND "STATO".stato_MODO_CW THEN
       "LINEARIZZA_POTENZA"(ingresso_in := #FWD_TMP_SS,
                            canale_in := 2,
                            tabella := "TABELLE_LINEARIZZAZIONE".tab_SS_CW,
                            uscita_out => "STATO".misura_FWD_SS);
   END_IF;
END_REGION
